(* Logix 5000 project; controller PLC_MCC1201_220AP1 vendor 1 type 14 code 164 rev 35.11; software revision 35.00; part 3 of 25 *)

   M212_M1_DR_MSF : MOTION_INSTRUCTION := (FLAGS := 570425344, DN := 1, STATUS := 2, STATE := 1); {access None}
   M212_M1_DR_MSO : MOTION_INSTRUCTION := (FLAGS := -1610612736, EN := 1, DN := 1, STATE := 1); {access None}
   M212_M1_DR_OUT_MAJ : MOTION_INSTRUCTION := (FLAGS := 570425344, DN := 1); {access None}
   M212_M1_DR_OUT_MAM : MOTION_INSTRUCTION := (FLAGS := 33554432); {access None}
   M212_M1_DR_OUT_MAR : MOTION_INSTRUCTION := (FLAGS := 33554432); {access None}
   M212_M1_DR_OUT_MAS : MOTION_INSTRUCTION := (FLAGS := -1442840576, EN := 1, DN := 1, PC := 1); {access None}
   M212_M1_DR_OUT_MCD : MOTION_INSTRUCTION := (FLAGS := 570425344, DN := 1); {access None}
   M212_M1_DR_OUT_MRP : MOTION_INSTRUCTION := (FLAGS := 33554432); {access None}
   M213_M1_DR : AXIS_CIP_DRIVE; {access Read Only}
   M213_M1_DR_IN_MAJ : MOTION_INSTRUCTION := (FLAGS := 570425344, DN := 1); {access None}
   M213_M1_DR_IN_MAM : MOTION_INSTRUCTION := (FLAGS := 33554432); {access None}
   M213_M1_DR_IN_MAR : MOTION_INSTRUCTION := (FLAGS := 33554432); {access None}
   M213_M1_DR_IN_MAS : MOTION_INSTRUCTION := (FLAGS := -1442840576, EN := 1, DN := 1, PC := 1); {access None}
   M213_M1_DR_IN_MCD : MOTION_INSTRUCTION := (FLAGS := 570425344, DN := 1); {access None}
   M213_M1_DR_IN_MRP : MOTION_INSTRUCTION := (FLAGS := 33554432); {access None}
   M213_M1_DR_MAFR : MOTION_INSTRUCTION := (FLAGS := 301989888, ER := 1, ERR := 11); {access None}
   M213_M1_DR_MDR : MOTION_INSTRUCTION := (FLAGS := -1845493760, EN := 1, ER := 1, ERR := 11); {access None}
   M213_M1_DR_MSF : MOTION_INSTRUCTION := (FLAGS := 570425344, DN := 1, STATUS := 2, STATE := 1); {access None}
   M213_M1_DR_MSO : MOTION_INSTRUCTION := (FLAGS := -1610612736, EN := 1, DN := 1, STATE := 1); {access None}
   M213_M1_DR_OUT_MAJ : MOTION_INSTRUCTION := (FLAGS := 570425344, DN := 1); {access None}
   M213_M1_DR_OUT_MAM : MOTION_INSTRUCTION := (FLAGS := 33554432); {access None}
   M213_M1_DR_OUT_MAR : MOTION_INSTRUCTION := (FLAGS := 33554432); {access None}
   M213_M1_DR_OUT_MAS : MOTION_INSTRUCTION := (FLAGS := -1442840576, EN := 1, DN := 1, PC := 1); {access None}
   M213_M1_DR_OUT_MCD : MOTION_INSTRUCTION := (FLAGS := 570425344, DN := 1); {access None}
   M213_M1_DR_OUT_MRP : MOTION_INSTRUCTION := (FLAGS := 33554432); {access None}
   M213A_M1_DR_IN_MAJ : MOTION_INSTRUCTION := (FLAGS := 570425344, DN := 1); {access None}
   M213A_M1_DR_IN_MAM : MOTION_INSTRUCTION := (FLAGS := 33554432); {access None}
   M213A_M1_DR_IN_MAR : MOTION_INSTRUCTION := (FLAGS := 33554432); {access None}
   M213A_M1_DR_IN_MAS : MOTION_INSTRUCTION := (FLAGS := -1442840576, EN := 1, DN := 1, PC := 1); {access None}
   M213A_M1_DR_IN_MCD : MOTION_INSTRUCTION := (FLAGS := 570425344, DN := 1); {access None}
   M213A_M1_DR_IN_MRP : MOTION_INSTRUCTION := (FLAGS := 33554432); {access None}
   M213A_M1_DR_MAFR : MOTION_INSTRUCTION := (FLAGS := 301989888, ER := 1, ERR := 11); {access None}
   M213A_M1_DR_MDR : MOTION_INSTRUCTION := (FLAGS := -1845493760, EN := 1, ER := 1, ERR := 11); {access None}
   M213A_M1_DR_MSF : MOTION_INSTRUCTION := (FLAGS := 570425344, DN := 1, STATUS := 2, STATE := 1); {access None}
   M213A_M1_DR_MSO : MOTION_INSTRUCTION := (FLAGS := -1610612736, EN := 1, DN := 1, STATE := 1); {access None}
   M213A_M1_DR_OUT_MAJ : MOTION_INSTRUCTION := (FLAGS := 570425344, DN := 1); {access None}
   M213A_M1_DR_OUT_MAM : MOTION_INSTRUCTION := (FLAGS := 33554432); {access None}
   M213A_M1_DR_OUT_MAR : MOTION_INSTRUCTION := (FLAGS := 33554432); {access None}
   M213A_M1_DR_OUT_MAS : MOTION_INSTRUCTION := (FLAGS := -1442840576, EN := 1, DN := 1, PC := 1); {access None}
   M213A_M1_DR_OUT_MCD : MOTION_INSTRUCTION := (FLAGS := 570425344, DN := 1); {access None}
   M213A_M1_DR_OUT_MRP : MOTION_INSTRUCTION := (FLAGS := 33554432); {access None}
   M213B_M1_DR_IN_MAJ : MOTION_INSTRUCTION := (FLAGS := 570425344, DN := 1); {access None}
   M213B_M1_DR_IN_MAM : MOTION_INSTRUCTION := (FLAGS := 33554432); {access None}
   M213B_M1_DR_IN_MAR : MOTION_INSTRUCTION := (FLAGS := 33554432); {access None}
   M213B_M1_DR_IN_MAS : MOTION_INSTRUCTION := (FLAGS := -1442840576, EN := 1, DN := 1, PC := 1); {access None}
   M213B_M1_DR_IN_MCD : MOTION_INSTRUCTION := (FLAGS := 570425344, DN := 1); {access None}
   M213B_M1_DR_IN_MRP : MOTION_INSTRUCTION := (FLAGS := 33554432); {access None}
   M213B_M1_DR_MAFR : MOTION_INSTRUCTION := (FLAGS := 301989888, ER := 1, ERR := 11); {access None}
   M213B_M1_DR_MDR : MOTION_INSTRUCTION := (FLAGS := -1845493760, EN := 1, ER := 1, ERR := 11); {access None}
   M213B_M1_DR_MSF : MOTION_INSTRUCTION := (FLAGS := 570425344, DN := 1, STATUS := 2, STATE := 1); {access None}
   M213B_M1_DR_MSO : MOTION_INSTRUCTION := (FLAGS := -1610612736, EN := 1, DN := 1, STATE := 1); {access None}
   M213B_M1_DR_OUT_MAJ : MOTION_INSTRUCTION := (FLAGS := 570425344, DN := 1); {access None}
   M213B_M1_DR_OUT_MAM : MOTION_INSTRUCTION := (FLAGS := 33554432); {access None}
   M213B_M1_DR_OUT_MAR : MOTION_INSTRUCTION := (FLAGS := 33554432); {access None}
   M213B_M1_DR_OUT_MAS : MOTION_INSTRUCTION := (FLAGS := -1442840576, EN := 1, DN := 1, PC := 1); {access None}
   M213B_M1_DR_OUT_MCD : MOTION_INSTRUCTION := (FLAGS := 570425344, DN := 1); {access None}
   M213B_M1_DR_OUT_MRP : MOTION_INSTRUCTION := (FLAGS := 33554432); {access None}
   M214_M1_DR : AXIS_CIP_DRIVE; {access Read Only}
   M214_M1_DR_IN_MAJ : MOTION_INSTRUCTION := (FLAGS := 570425344, DN := 1); {access None}
   M214_M1_DR_IN_MAM : MOTION_INSTRUCTION := (FLAGS := 33554432); {access None}
   M214_M1_DR_IN_MAR : MOTION_INSTRUCTION := (FLAGS := 33554432); {access None}
   M214_M1_DR_IN_MAS : MOTION_INSTRUCTION := (FLAGS := -1442840576, EN := 1, DN := 1, PC := 1); {access None}
   M214_M1_DR_IN_MCD : MOTION_INSTRUCTION := (FLAGS := 570425344, DN := 1); {access None}
   M214_M1_DR_IN_MRP : MOTION_INSTRUCTION := (FLAGS := 33554432); {access None}
   M214_M1_DR_MAFR : MOTION_INSTRUCTION := (FLAGS := 301989888, ER := 1, ERR := 11); {access None}
   M214_M1_DR_MDR : MOTION_INSTRUCTION := (FLAGS := -1845493760, EN := 1, ER := 1, ERR := 11); {access None}
   M214_M1_DR_MSF : MOTION_INSTRUCTION := (FLAGS := 570425344, DN := 1, STATUS := 2, STATE := 1); {access None}
   M214_M1_DR_MSO : MOTION_INSTRUCTION := (FLAGS := -1610612736, EN := 1, DN := 1, STATE := 1); {access None}
   M214_M1_DR_OUT_MAJ : MOTION_INSTRUCTION := (FLAGS := 570425344, DN := 1); {access None}
   M214_M1_DR_OUT_MAM : MOTION_INSTRUCTION := (FLAGS := 33554432); {access None}
   M214_M1_DR_OUT_MAR : MOTION_INSTRUCTION := (FLAGS := 33554432); {access None}
   M214_M1_DR_OUT_MAS : MOTION_INSTRUCTION := (FLAGS := -1442840576, EN := 1, DN := 1, PC := 1); {access None}
   M214_M1_DR_OUT_MCD : MOTION_INSTRUCTION := (FLAGS := 570425344, DN := 1); {access None}
   M214_M1_DR_OUT_MRP : MOTION_INSTRUCTION := (FLAGS := 33554432); {access None}
   M215_M1_DR : AXIS_CIP_DRIVE; {access Read Only}
   M215_M1_DR_IN_MAJ : MOTION_INSTRUCTION := (FLAGS := 570425344, DN := 1); {access None}
   M215_M1_DR_IN_MAM : MOTION_INSTRUCTION := (FLAGS := 33554432); {access None}
   M215_M1_DR_IN_MAR : MOTION_INSTRUCTION := (FLAGS := 33554432); {access None}
   M215_M1_DR_IN_MAS : MOTION_INSTRUCTION := (FLAGS := -1442840576, EN := 1, DN := 1, PC := 1); {access None}
   M215_M1_DR_IN_MCD : MOTION_INSTRUCTION := (FLAGS := 570425344, DN := 1); {access None}
   M215_M1_DR_IN_MRP : MOTION_INSTRUCTION := (FLAGS := 33554432); {access None}
   M215_M1_DR_MAFR : MOTION_INSTRUCTION := (FLAGS := 301989888, ER := 1, ERR := 11); {access None}
   M215_M1_DR_MDR : MOTION_INSTRUCTION := (FLAGS := -1845493760, EN := 1, ER := 1, ERR := 11); {access None}
   M215_M1_DR_MSF : MOTION_INSTRUCTION := (FLAGS := 570425344, DN := 1, STATUS := 2, STATE := 1); {access None}
   M215_M1_DR_MSO : MOTION_INSTRUCTION := (FLAGS := -1610612736, EN := 1, DN := 1, STATE := 1); {access None}
   M215_M1_DR_OUT_MAJ : MOTION_INSTRUCTION := (FLAGS := 570425344, DN := 1); {access None}
   M215_M1_DR_OUT_MAM : MOTION_INSTRUCTION := (FLAGS := 33554432); {access None}
   M215_M1_DR_OUT_MAR : MOTION_INSTRUCTION := (FLAGS := 33554432); {access None}
   M215_M1_DR_OUT_MAS : MOTION_INSTRUCTION := (FLAGS := -1442840576, EN := 1, DN := 1, PC := 1); {access None}
   M215_M1_DR_OUT_MCD : MOTION_INSTRUCTION := (FLAGS := 570425344, DN := 1); {access None}
   M215_M1_DR_OUT_MRP : MOTION_INSTRUCTION := (FLAGS := 33554432); {access None}
   M216_M1_DR : AXIS_CIP_DRIVE; {access Read Only}
   M216_M1_DR_IN_MAJ : MOTION_INSTRUCTION := (FLAGS := 570425344, DN := 1); {access None}
   M216_M1_DR_IN_MAM : MOTION_INSTRUCTION := (FLAGS := 33554432); {access None}
   M216_M1_DR_IN_MAR : MOTION_INSTRUCTION := (FLAGS := 33554432); {access None}
   M216_M1_DR_IN_MAS : MOTION_INSTRUCTION := (FLAGS := -1442840576, EN := 1, DN := 1, PC := 1); {access None}
   M216_M1_DR_IN_MCD : MOTION_INSTRUCTION := (FLAGS := 570425344, DN := 1); {access None}
   M216_M1_DR_IN_MRP : MOTION_INSTRUCTION := (FLAGS := 33554432); {access None}
   M216_M1_DR_MAFR : MOTION_INSTRUCTION := (FLAGS := 301989888, ER := 1, ERR := 11); {access None}
   M216_M1_DR_MDR : MOTION_INSTRUCTION := (FLAGS := -1845493760, EN := 1, ER := 1, ERR := 11); {access None}
   M216_M1_DR_MSF : MOTION_INSTRUCTION := (FLAGS := 570425344, DN := 1, STATUS := 2, STATE := 1); {access None}
   M216_M1_DR_MSO : MOTION_INSTRUCTION := (FLAGS := -1610612736, EN := 1, DN := 1, STATE := 1); {access None}
   M216_M1_DR_OUT_MAJ : MOTION_INSTRUCTION := (FLAGS := 570425344, DN := 1); {access None}
   M216_M1_DR_OUT_MAM : MOTION_INSTRUCTION := (FLAGS := 33554432); {access None}
   M216_M1_DR_OUT_MAR : MOTION_INSTRUCTION := (FLAGS := 33554432); {access None}
   M216_M1_DR_OUT_MAS : MOTION_INSTRUCTION := (FLAGS := -1442840576, EN := 1, DN := 1, PC := 1); {access None}
   M216_M1_DR_OUT_MCD : MOTION_INSTRUCTION := (FLAGS := 570425344, DN := 1); {access None}
   M216_M1_DR_OUT_MRP : MOTION_INSTRUCTION := (FLAGS := 33554432); {access None}
   M217_M1_DR : AXIS_CIP_DRIVE; {access Read Only}
   M217_M1_DR_IN_MAJ : MOTION_INSTRUCTION := (FLAGS := 570425344, DN := 1); {access None}
   M217_M1_DR_IN_MAM : MOTION_INSTRUCTION := (FLAGS := 33554432); {access None}
   M217_M1_DR_IN_MAR : MOTION_INSTRUCTION := (FLAGS := 33554432); {access None}
   M217_M1_DR_IN_MAS : MOTION_INSTRUCTION := (FLAGS := -1442840576, EN := 1, DN := 1, PC := 1); {access None}
   M217_M1_DR_IN_MCD : MOTION_INSTRUCTION := (FLAGS := 570425344, DN := 1); {access None}
   M217_M1_DR_IN_MRP : MOTION_INSTRUCTION := (FLAGS := 33554432); {access None}
   M217_M1_DR_MAFR : MOTION_INSTRUCTION := (FLAGS := 301989888, ER := 1, ERR := 11); {access None}
   M217_M1_DR_MDR : MOTION_INSTRUCTION := (FLAGS := -1845493760, EN := 1, ER := 1, ERR := 11); {access None}
   M217_M1_DR_MSF : MOTION_INSTRUCTION := (FLAGS := 570425344, DN := 1, STATUS := 2, STATE := 1); {access None}
   M217_M1_DR_MSO : MOTION_INSTRUCTION := (FLAGS := -1610612736, EN := 1, DN := 1, STATE := 1); {access None}
   M217_M1_DR_OUT_MAJ : MOTION_INSTRUCTION := (FLAGS := 570425344, DN := 1); {access None}
   M217_M1_DR_OUT_MAM : MOTION_INSTRUCTION := (FLAGS := 33554432); {access None}
   M217_M1_DR_OUT_MAR : MOTION_INSTRUCTION := (FLAGS := 33554432); {access None}
   M217_M1_DR_OUT_MAS : MOTION_INSTRUCTION := (FLAGS := -1442840576, EN := 1, DN := 1, PC := 1); {access None}
   M217_M1_DR_OUT_MCD : MOTION_INSTRUCTION := (FLAGS := 570425344, DN := 1); {access None}
   M217_M1_DR_OUT_MRP : MOTION_INSTRUCTION := (FLAGS := 33554432); {access None}
   M218_M1_DR : AXIS_CIP_DRIVE; {access Read Only}
   M218_M1_DR_IN_MAJ : MOTION_INSTRUCTION := (FLAGS := 570425344, DN := 1); {access None}
   M218_M1_DR_IN_MAM : MOTION_INSTRUCTION := (FLAGS := 33554432); {access None}
   M218_M1_DR_IN_MAR : MOTION_INSTRUCTION := (FLAGS := 33554432); {access None}
   M218_M1_DR_IN_MAS : MOTION_INSTRUCTION := (FLAGS := -1442840576, EN := 1, DN := 1, PC := 1); {access None}
   M218_M1_DR_IN_MCD : MOTION_INSTRUCTION := (FLAGS := 570425344, DN := 1); {access None}
   M218_M1_DR_IN_MRP : MOTION_INSTRUCTION := (FLAGS := 33554432); {access None}
   M218_M1_DR_MAFR : MOTION_INSTRUCTION := (FLAGS := 301989888, ER := 1, ERR := 11); {access None}
   M218_M1_DR_MDR : MOTION_INSTRUCTION := (FLAGS := -1845493760, EN := 1, ER := 1, ERR := 11); {access None}
   M218_M1_DR_MSF : MOTION_INSTRUCTION := (FLAGS := 570425344, DN := 1, STATUS := 2, STATE := 1); {access None}
   M218_M1_DR_MSO : MOTION_INSTRUCTION := (FLAGS := -1610612736, EN := 1, DN := 1, STATE := 1); {access None}
   M218_M1_DR_OUT_MAJ : MOTION_INSTRUCTION := (FLAGS := 570425344, DN := 1); {access None}
   M218_M1_DR_OUT_MAM : MOTION_INSTRUCTION := (FLAGS := 33554432); {access None}
   M218_M1_DR_OUT_MAR : MOTION_INSTRUCTION := (FLAGS := 33554432); {access None}
   M218_M1_DR_OUT_MAS : MOTION_INSTRUCTION := (FLAGS := -1442840576, EN := 1, DN := 1, PC := 1); {access None}
   M218_M1_DR_OUT_MCD : MOTION_INSTRUCTION := (FLAGS := 570425344, DN := 1); {access None}
   M218_M1_DR_OUT_MRP : MOTION_INSTRUCTION := (FLAGS := 33554432); {access None}
   M219_M1_DR : AXIS_CIP_DRIVE; {access Read Only}
   M219_M1_DR_IN_MAJ : MOTION_INSTRUCTION := (FLAGS := 570425344, DN := 1); {access None}
   M219_M1_DR_IN_MAM : MOTION_INSTRUCTION := (FLAGS := 33554432); {access None}
   M219_M1_DR_IN_MAR : MOTION_INSTRUCTION := (FLAGS := 33554432); {access None}
   M219_M1_DR_IN_MAS : MOTION_INSTRUCTION := (FLAGS := -1442840576, EN := 1, DN := 1, PC := 1); {access None}
   M219_M1_DR_IN_MCD : MOTION_INSTRUCTION := (FLAGS := 570425344, DN := 1); {access None}
   M219_M1_DR_IN_MRP : MOTION_INSTRUCTION := (FLAGS := 33554432); {access None}
   M219_M1_DR_MAFR : MOTION_INSTRUCTION := (FLAGS := 301989888, ER := 1, ERR := 11); {access None}
   M219_M1_DR_MDR : MOTION_INSTRUCTION := (FLAGS := -1845493760, EN := 1, ER := 1, ERR := 11); {access None}
   M219_M1_DR_MSF : MOTION_INSTRUCTION := (FLAGS := 570425344, DN := 1, STATUS := 2, STATE := 1); {access None}
   M219_M1_DR_MSO : MOTION_INSTRUCTION := (FLAGS := -1610612736, EN := 1, DN := 1, STATE := 1); {access None}
   M219_M1_DR_OUT_MAJ : MOTION_INSTRUCTION := (FLAGS := 570425344, DN := 1); {access None}
   M219_M1_DR_OUT_MAM : MOTION_INSTRUCTION := (FLAGS := 33554432); {access None}
   M219_M1_DR_OUT_MAR : MOTION_INSTRUCTION := (FLAGS := 33554432); {access None}
   M219_M1_DR_OUT_MAS : MOTION_INSTRUCTION := (FLAGS := -1442840576, EN := 1, DN := 1, PC := 1); {access None}
   M219_M1_DR_OUT_MCD : MOTION_INSTRUCTION := (FLAGS := 570425344, DN := 1); {access None}
   M219_M1_DR_OUT_MRP : MOTION_INSTRUCTION := (FLAGS := 33554432); {access None}
   M220_M1_DR : AXIS_CIP_DRIVE; {access Read Only}
   M220_M1_DR_IN_MAJ : MOTION_INSTRUCTION := (FLAGS := 570425344, DN := 1); {access None}
   M220_M1_DR_IN_MAM : MOTION_INSTRUCTION := (FLAGS := 33554432); {access None}
   M220_M1_DR_IN_MAR : MOTION_INSTRUCTION := (FLAGS := 33554432); {access None}
   M220_M1_DR_IN_MAS : MOTION_INSTRUCTION := (FLAGS := -1442840576, EN := 1, DN := 1, PC := 1); {access None}
   M220_M1_DR_IN_MCD : MOTION_INSTRUCTION := (FLAGS := 570425344, DN := 1); {access None}
   M220_M1_DR_IN_MRP : MOTION_INSTRUCTION := (FLAGS := 33554432); {access None}
   M220_M1_DR_MAFR : MOTION_INSTRUCTION := (FLAGS := 301989888, ER := 1, ERR := 11); {access None}
   M220_M1_DR_MDR : MOTION_INSTRUCTION := (FLAGS := -1845493760, EN := 1, ER := 1, ERR := 11); {access None}
   M220_M1_DR_MSF : MOTION_INSTRUCTION := (FLAGS := 570425344, DN := 1, STATUS := 2, STATE := 1); {access None}
   M220_M1_DR_MSO : MOTION_INSTRUCTION := (FLAGS := -1610612736, EN := 1, DN := 1, STATE := 1); {access None}
   M220_M1_DR_OUT_MAJ : MOTION_INSTRUCTION := (FLAGS := 570425344, DN := 1); {access None}
   M220_M1_DR_OUT_MAM : MOTION_INSTRUCTION := (FLAGS := 33554432); {access None}
   M220_M1_DR_OUT_MAR : MOTION_INSTRUCTION := (FLAGS := 33554432); {access None}
   M220_M1_DR_OUT_MAS : MOTION_INSTRUCTION := (FLAGS := -1442840576, EN := 1, DN := 1, PC := 1); {access None}
   M220_M1_DR_OUT_MCD : MOTION_INSTRUCTION := (FLAGS := 570425344, DN := 1); {access None}
   M220_M1_DR_OUT_MRP : MOTION_INSTRUCTION := (FLAGS := 33554432); {access None}
   M225 : MAC_EMERGENCYXCUT := (ST_xConditionOKAccessArea := 1, ST_xSelectorManualMode := 1, ST_xManualModeSelection := 1, ST_xManualModeAccepted := 1, ST_xDistanceBetweenCutOK := 1, ST_xConditionOKStopCycle := 1, ST_xConditionOKSemiautoMode := 1, ST_xConditionOKManualMode := 1, ST_xBreakerCutRequest := 1, OUTPUT_xMachineOutOfOrder := 1, OUTPUT_xAreaSafetyOn := 1, OUTPUT_xStopCut := 1, AUX_dDistanceFTCHead := 6050, AUX_dBridgeAngle := 80000, AUX_dManualSpeed_mm_min := 10000, AUX_dRiseReactionTime_ms := 50, AUX_dDescentReactionTime_ms := 1000, AUX_dBackwardFastSpeed_mm_min := 120000, AUX_dBackwardSlowSpeed_mm_min := 90000, AUX_dCarriageFinalPosition_cmm := 400000, AUX_dMinimumStripeLength := 100000, AUX_dMaximumStripeLength := 300000, AUX_dLastCutValue := -268936272, AUX_dLastCutValueStored := -268936272, AUX_dForwardTimeoutTime_ms := 2147483647, AUX_dReturnSpeed_mm_min := 90000, AUX_dReqSpeed_mm_min := 10000, AUX_dStartControlPhotocellPos_dmm := -36050, AUX_dTimeFTCToHead_ms := 36300000, AUX_dTimeDelayToDescent_ms := 36299800, AUX_dTimeAdvanceToRise_ms := 36293450, AUX_dTimeDelayToLubrication_ms := 36300000, OSR_xConditionNotOKToCut := 1, AUX_tmOFF_DriveEnable.PRE := 100, AUX_tmOFF_DriveEnable.ACC := 100, AUX_tmOFF_AreaSafetyOK.PRE := 2000, AUX_tmOFF_AreaSafetyOK.ACC := 2000, AUX_tmON_FdbkError.PRE := 2000, AUX_tmON_TimeoutHome.PRE := 90000, AUX_tmON_TimeoutFW.PRE := 120000, AUX_tmON_TimeoutBW.PRE := 90000, AUX_tmOFF_LowerHeadNotAllowed.PRE := 200, AUX_tmOFF_LowerHeadNotAllowed.ACC := 200, AUX_tmOFF_AdvanceTimeToRise.PRE := 171, AUX_tmOFF_AdvanceTimeToRise.ACC := 171, AUX_tmON_DelayTimeLubrication.PRE := 221, AUX_tmON_DelayTimeLubrication.ACC := 221, AUX_tmON_TimeoutHeadPosition.PRE := 90000, CONST_dAcceleration_m_s2 := 3, CONST_dDeceleration_m_s2 := 3); {access None}
   M225_ALM : MAC_EMERGENCYXCUT_ALM; {access Read Only}
        .rgxStoppingFaults[0].4   // A120KE1.Area safety
        .rgxStoppingFaults[0].8   // A57AZ1.Timeout move backward
        .rgxStoppingFaults[0].2   // A57AZ1.Drive error
        .rgxStoppingFaults[0].9   // A57AZ1.Timeout home position (A121SQ1)
        .rgxStoppingFaults[0].1   // A207BT2.Motor thermal probe
        .rgxFaults[0].0   // A57QM1.Protection traslation
        .rgxFaults[0].1   // A57QM2.Protection fan rotation
        .rgdCodeAlarm[0].0   // A63AZ1.Code alarm
        .rgxStoppingFaults[0].7   // A57AZ1.Timeout move forward
        .rgxStoppingFaults[0].11   // A207SP1.Compressed air failure
        .rgxStoppingFaults[0].10   // A208SQ1.Error position cutting head
        .rgxStoppingFaults[0].5   // A121SQ1.Forward Overstroke
        .rgxStoppingFaults[0].6   // A121SQ2.Backward Overstroke
        .rgxStoppingFaults[0].3   // A57AZ1.Traslation feedback
        .rgxStoppingFaults[0].0   // A57QS1.Safety motor sectioning
   M225_HMR : MAC_EMERGENCYXCUT_HMR := (dMode := 1, dStatus := 1, dZoneStatus := 2, dDistanceFromSnaproll_cmm := 5050000, rHeadUsage_km := 0.0004); {access Read Only}
   M225_HMW : MAC_EMERGENCYXCUT_HMW := (dLowerHeadDelayTime_ms := 800, dRiseHeadAdvanceTime_ms := 6500, dCulletStripeLength_cmm := 220000, dDistanceFromSnaproll_cmm := 5030000);
   M225_IN_MOTION : MAC_EMERGENCYXCUT_IN_MOTION; {access None}
   M225_M1_DR : AXIS_CIP_DRIVE; {access Read Only}
   M225_M1_DR_IN_MAJ : MOTION_INSTRUCTION := (FLAGS := 570425344, DN := 1); {access None}
   M225_M1_DR_IN_MAM : MOTION_INSTRUCTION := (FLAGS := 33554432); {access None}
   M225_M1_DR_IN_MAR : MOTION_INSTRUCTION := (FLAGS := 33554432); {access None}
   M225_M1_DR_IN_MAS : MOTION_INSTRUCTION := (FLAGS := -1442840576, EN := 1, DN := 1, PC := 1); {access None}
   M225_M1_DR_IN_MCD : MOTION_INSTRUCTION := (FLAGS := 570425344, DN := 1); {access None}
   M225_M1_DR_IN_MRP : MOTION_INSTRUCTION := (FLAGS := 33554432); {access None}
   M225_M1_DR_MAFR : MOTION_INSTRUCTION := (FLAGS := 301989888, ER := 1, ERR := 11); {access None}
   M225_M1_DR_MDR : MOTION_INSTRUCTION := (FLAGS := -1845493760, EN := 1, ER := 1, ERR := 11); {access None}
   M225_M1_DR_MSF : MOTION_INSTRUCTION := (FLAGS := 570425344, DN := 1, STATUS := 2, STATE := 1); {access None}
   M225_M1_DR_MSO : MOTION_INSTRUCTION := (FLAGS := -1610612736, EN := 1, DN := 1, STATE := 1); {access None}
   M225_M1_DR_OUT_MAJ : MOTION_INSTRUCTION := (FLAGS := 570425344, DN := 1); {access None}
   M225_M1_DR_OUT_MAM : MOTION_INSTRUCTION := (FLAGS := 33554432); {access None}
   M225_M1_DR_OUT_MAR : MOTION_INSTRUCTION := (FLAGS := 33554432); {access None}
   M225_M1_DR_OUT_MAS : MOTION_INSTRUCTION := (FLAGS := -1442840576, EN := 1, DN := 1, PC := 1); {access None}
   M225_M1_DR_OUT_MCD : MOTION_INSTRUCTION := (FLAGS := 570425344, DN := 1); {access None}
   M225_M1_DR_OUT_MRP : MOTION_INSTRUCTION := (FLAGS := 33554432); {access None}
   M225_OUT_MOTION : MAC_EMERGENCYXCUT_OUT_MOTION := (DR_MSO.FLAGS := 33554432, DR_MSF.FLAGS := -1577058304, DR_MSF.EN := 1, DR_MSF.DN := 1, DR_MSF.STATUS := 2, DR_MSF.STATE := 1, DR_MASR.FLAGS := 33554432, DR_MAJ.FLAGS := 33554432, DR_MAM.FLAGS := 33554432, DR_MAS.FLAGS := -1442840576, DR_MAS.EN := 1, DR_MAS.DN := 1, DR_MAS.PC := 1, DR_MAH.FLAGS := 33554432); {access None}
   M225S_AOI_AccessArea : STRUCT_AccessArea := (tAccess[0].tHMR.dStatusAccessArea := 4, tAccess[0].tSTC.IN_xConditionOkAccessArea := 1, tAccess[0].tSTC.OUT_xSafetyAreaIntervened := 1, tAccess[1].tHMR.dStatusAccessArea := 4, tAccess[1].tSTC.OUT_xSafetyAreaIntervened := 1);
   M2xx_CONVEYOR : MAC_CONVEYOR[20] := ([0].AUX_tmOFFRetainDriveEnable.PRE := 1000, [0].AUX_tmOFFRetainDriveEnable.ACC := 1000, [0].AUX_tmONRotfeedBackAlarm.PRE := 2000, [0].AUX_tmONDriveReadyAlarm.PRE := 1000, [0].AUX_rAcceleration_m_s2 := 0.25, [0].AUX_rDeceleration_m_s2 := 0.25, [0].AUX_dReqSpeed_mm_min := 6807, [0].AUX_dRealSpeed_mm_min := 6807, [1].AUX_tmOFFRetainDriveEnable.PRE := 1000, [1].AUX_tmOFFRetainDriveEnable.ACC := 1000, [1].AUX_tmONDriveReadyAlarm.PRE := 1000, [1].AUX_rAcceleration_m_s2 := 0.25, [1].AUX_rDeceleration_m_s2 := 0.25, [1].AUX_dReqSpeed_mm_min := 6807, [1].AUX_dRealSpeed_mm_min := 6807, [2].INPUT_xProtectionFan := 1, [2].AUX_tmOFFRetainDriveEnable.PRE := 1000, [2].AUX_tmOFFRetainDriveEnable.ACC := 1000, [2].AUX_tmONDriveReadyAlarm.PRE := 1000, [2].AUX_rAcceleration_m_s2 := 0.25, [2].AUX_rDeceleration_m_s2 := 0.25, [2].AUX_dReqSpeed_mm_min := 6807, [2].AUX_dRealSpeed_mm_min := 6807, [3].INPUT_xProtectionFan := 1, [3].AUX_tmOFFRetainDriveEnable.PRE := 1000, [3].AUX_tmOFFRetainDriveEnable.ACC := 1000, [3].AUX_tmONDriveReadyAlarm.PRE := 1000, [3].AUX_rAcceleration_m_s2 := 0.25, [3].AUX_rDeceleration_m_s2 := 0.25, [3].AUX_dReqSpeed_mm_min := 6807, [3].AUX_dRealSpeed_mm_min := 6807, [4].INPUT_xProtectionFan := 1, [4].AUX_tmOFFRetainDriveEnable.PRE := 1000, [4].AUX_tmOFFRetainDriveEnable.ACC := 1000, [4].AUX_tmONDriveReadyAlarm.PRE := 1000, [4].AUX_rAcceleration_m_s2 := 0.25, [4].AUX_rDeceleration_m_s2 := 0.25, [4].AUX_dReqSpeed_mm_min := 6807, [4].AUX_dRealSpeed_mm_min := 6807, [5].ST_xStoppingFaults := 1, [5].INPUT_xProtectionFan := 1, [5].AUX_tmOFFRetainDriveEnable.PRE := 1000, [5].AUX_tmOFFRetainDriveEnable.ACC := 1000, [5].AUX_tmONDriveReadyAlarm.PRE := 1000, [5].AUX_rAcceleration_m_s2 := 0.25, [5].AUX_rDeceleration_m_s2 := 0.25, [5].AUX_dReqSpeed_mm_min := 6807, [5].AUX_dRealSpeed_mm_min := 6807, [6].ST_xStoppingFaults := 1, [6].INPUT_xProtectionFan := 1, [6].AUX_tmOFFRetainDriveEnable.PRE := 1000, [6].AUX_tmOFFRetainDriveEnable.ACC := 1000, [6].AUX_tmONDriveReadyAlarm.PRE := 1000, [6].AUX_rAcceleration_m_s2 := 0.25, [6].AUX_rDeceleration_m_s2 := 0.25, [6].AUX_dReqSpeed_mm_min := 6807, [6].AUX_dRealSpeed_mm_min := 6807, [7].ST_xStoppingFaults := 1, [7].INPUT_xProtectionFan := 1, [7].AUX_tmOFFRetainDriveEnable.PRE := 1000,
        [7].AUX_tmOFFRetainDriveEnable.ACC := 1000, [7].AUX_tmONDriveReadyAlarm.PRE := 1000, [7].AUX_rAcceleration_m_s2 := 0.25, [7].AUX_rDeceleration_m_s2 := 0.25, [7].AUX_dReqSpeed_mm_min := 6807, [7].AUX_dRealSpeed_mm_min := 6807, [8].ST_xStoppingFaults := 1, [8].INPUT_xProtectionFan := 1, [8].AUX_tmOFFRetainDriveEnable.PRE := 1000, [8].AUX_tmOFFRetainDriveEnable.ACC := 1000, [8].AUX_tmONDriveReadyAlarm.PRE := 1000, [8].AUX_rAcceleration_m_s2 := 0.25, [8].AUX_rDeceleration_m_s2 := 0.25, [8].AUX_dReqSpeed_mm_min := 6807, [8].AUX_dRealSpeed_mm_min := 6807, [9].ST_xStoppingFaults := 1, [9].INPUT_xProtectionFan := 1, [9].AUX_tmOFFRetainDriveEnable.PRE := 1000, [9].AUX_tmOFFRetainDriveEnable.ACC := 1000, [9].AUX_tmONDriveReadyAlarm.PRE := 1000, [9].AUX_rAcceleration_m_s2 := 0.25, [9].AUX_rDeceleration_m_s2 := 0.25, [9].AUX_dReqSpeed_mm_min := 6807, [9].AUX_dRealSpeed_mm_min := 6807, [10].ST_xStoppingFaults := 1, [10].INPUT_xProtectionFan := 1, [10].AUX_tmOFFRetainDriveEnable.PRE := 1000, [10].AUX_tmOFFRetainDriveEnable.ACC := 1000, [10].AUX_tmONDriveReadyAlarm.PRE := 1000, [10].AUX_rAcceleration_m_s2 := 0.25, [10].AUX_rDeceleration_m_s2 := 0.25, [10].AUX_dReqSpeed_mm_min := 6807, [10].AUX_dRealSpeed_mm_min := 6807, [11].INPUT_xProtectionFan := 1, [11].AUX_tmOFFRetainDriveEnable.PRE := 1000, [11].AUX_tmOFFRetainDriveEnable.ACC := 1000, [11].AUX_tmONDriveReadyAlarm.PRE := 1000, [11].AUX_rAcceleration_m_s2 := 0.25, [11].AUX_rDeceleration_m_s2 := 0.25, [11].AUX_dReqSpeed_mm_min := 6807, [11].AUX_dRealSpeed_mm_min := 6807, [12].INPUT_xProtectionFan := 1, [12].AUX_tmOFFRetainDriveEnable.PRE := 1000, [12].AUX_tmOFFRetainDriveEnable.ACC := 1000, [12].AUX_dReqSpeed_mm_min := 6807, [12].AUX_dRealSpeed_mm_min := 6807, [13].INPUT_xProtectionFan := 1, [13].AUX_tmOFFRetainDriveEnable.PRE := 1000, [13].AUX_tmOFFRetainDriveEnable.ACC := 1000, [13].AUX_dReqSpeed_mm_min := 6807, [13].AUX_dRealSpeed_mm_min := 6807, [14].INPUT_xProtectionFan := 1, [14].AUX_tmOFFRetainDriveEnable.PRE := 1000, [14].AUX_tmOFFRetainDriveEnable.ACC := 1000, [14].AUX_dReqSpeed_mm_min := 6807, [14].AUX_dRealSpeed_mm_min := 6807, [15].INPUT_xProtectionFan := 1, [15].AUX_tmOFFRetainDriveEnable.PRE := 1000, [15].AUX_tmOFFRetainDriveEnable.ACC := 1000, [15].AUX_dReqSpeed_mm_min := 6807,
        [15].AUX_dRealSpeed_mm_min := 6807, [16].INPUT_xProtectionFan := 1, [16].AUX_tmOFFRetainDriveEnable.PRE := 1000, [16].AUX_tmOFFRetainDriveEnable.ACC := 1000, [16].AUX_dReqSpeed_mm_min := 6807, [16].AUX_dRealSpeed_mm_min := 6807, [17].INPUT_xProtectionFan := 1, [17].AUX_tmOFFRetainDriveEnable.PRE := 1000, [17].AUX_tmOFFRetainDriveEnable.ACC := 1000, [17].AUX_dReqSpeed_mm_min := 6807, [17].AUX_dRealSpeed_mm_min := 6807, [18].INPUT_xProtectionFan := 1, [18].AUX_tmOFFRetainDriveEnable.PRE := 1000, [18].AUX_tmOFFRetainDriveEnable.ACC := 1000, [18].AUX_dReqSpeed_mm_min := 6807, [18].AUX_dRealSpeed_mm_min := 6807, [19].INPUT_xProtectionFan := 1, [19].AUX_tmOFFRetainDriveEnable.PRE := 1000, [19].AUX_tmOFFRetainDriveEnable.ACC := 1000, [19].AUX_dReqSpeed_mm_min := 6807, [19].AUX_dRealSpeed_mm_min := 6807); {access None}
        [0]   // M202
        [10]   // M213
        [1]   // M203
        [2]   // M204
        [3]   // M206
        [4]   // M207
        [5]   // M208
        [6]   // M209
        [7]   // M210
        [8]   // M211
        [9]   // M212
        [11]   // M214
        [12]   // M215
        [13]   // M216
        [14]   // M217
        [15]   // M218
        [19]   // M301M2
        [18]   // M301M1
        [16]   // M219
        [17]   // M220
   M2xx_CONVEYOR_ALM : MAC_CONVEYOR_ALM[20] := ([5].rgxStoppingFaults[0] := 16, [6].rgxStoppingFaults[0] := 16, [7].rgxStoppingFaults[0] := 16, [8].rgxStoppingFaults[0] := 16, [9].rgxStoppingFaults[0] := 16, [10].rgxStoppingFaults[0] := 16); {access Read Only}
        [0]   // M202
        [0].rgxStoppingFaults[0].2   // A53AZ1.Drive error
        [2].rgxStoppingFaults[0].2   // A55AZ1.Drive error
        [1].rgxStoppingFaults[0].2   // A54AZ1.Drive error
        [0].rgdCodeAlarm[0].0   // AZ.Drive error code
        [0].rgxFaults[0].0   // QM.Protection fan rotation
        [10]   // M213
        [11]   // M214
        [1]   // M203
        [2]   // M204
        [3]   // M206
        [4]   // M207
        [5]   // M208
        [6]   // M209
        [7]   // M210
        [8]   // M211
        [9]   // M212
        [17]   // M220
        [18]   // M301M1
        [16]   // M219
        [15]   // M218
        [14]   // M217
        [13]   // M216
        [12]   // M215
        [19]   // M301M2
        [0].rgxStoppingFaults[0].1   // A206BT1.Motor thermal probe
        [1].rgxStoppingFaults[0].1   // A206BT2.Motor thermal probe
        [1].rgxStoppingFaults[0].3   // A54AZ1.Rotation feedback
        [0].rgxStoppingFaults[0].0   // A53QS1.Local safety switch
        [0].rgxStoppingFaults[0].4   // A53AZ1.Drive not ready
        [1].rgxStoppingFaults[0].0   // A54QS1.Local safety switch
        [0].rgxStoppingFaults[0].3   // A53AZ1.Rotation feedback
        [1].rgxStoppingFaults[0].4   // A54AZ1.Drive not ready
        [2].rgxStoppingFaults[0].0   // A55QS1.Local safety switch
        [2].rgxStoppingFaults[0].1   // A207BT1.Motor thermal probe
        [2].rgxStoppingFaults[0].3   // A55AZ1.Rotation feedback
        [2].rgxStoppingFaults[0].4   // A55AZ1.Drive not ready
        [3].rgxStoppingFaults[0].0   // A61QS1.Local safety switch
        [3].rgxStoppingFaults[0].1   // A209BT1.Motor thermal probe
        [3].rgxStoppingFaults[0].2   // A61AZ1.Drive error
        [3].rgxStoppingFaults[0].3   // A61AZ1.Rotation feedback
        [3].rgxStoppingFaults[0].4   // A61AZ1.Drive not ready
        [4].rgxStoppingFaults[0].0   // A62QS1.Local safety switch
        [5].rgxStoppingFaults[0].0   // A63QS1.Local safety switch
        [6].rgxStoppingFaults[0].0   // A64QS1.Local safety switch
        [7].rgxStoppingFaults[0].0   // A65QS1.Local safety switch
        [8].rgxStoppingFaults[0].0   // A66QS1.Local safety switch
        [9].rgxStoppingFaults[0].0   // A67QS1.Local safety switch
        [10].rgxStoppingFaults[0].0   // A68QS1.Local safety switch
        [11].rgxStoppingFaults[0].0   // A69QS1.Local safety switch
        [12].rgxStoppingFaults[0].0   // A70QS1.Local safety switch
        [13].rgxStoppingFaults[0].0   // A71QS1.Local safety switch
        [14].rgxStoppingFaults[0].0   // A72QS1.Local safety switch
        [15].rgxStoppingFaults[0].0   // A73QS1.Local safety switch
        [16].rgxStoppingFaults[0].0   // A74QS1.Local safety switch
        [17].rgxStoppingFaults[0].0   // A77QS1.Local safety switch
        [4].rgxStoppingFaults[0].1   // A209BT2.Motor thermal probe
        [5].rgxStoppingFaults[0].1   // A209BT3.Motor thermal probe
        [6].rgxStoppingFaults[0].1   // A209BT4.Motor thermal probe
        [7].rgxStoppingFaults[0].1   // A209BT5.Motor thermal probe
        [8].rgxStoppingFaults[0].1   // A209BT6.Motor thermal probe
        [9].rgxStoppingFaults[0].1   // A209BT7.Motor thermal probe
        [10].rgxStoppingFaults[0].1   // A209BT8.Motor thermal probe
        [11].rgxStoppingFaults[0].1   // A210BT1.Motor thermal probe
        [12].rgxStoppingFaults[0].1   // A210BT2.Motor thermal probe
        [13].rgxStoppingFaults[0].1   // A210BT3.Motor thermal probe
        [14].rgxStoppingFaults[0].1   // A210BT4.Motor thermal probe
        [15].rgxStoppingFaults[0].1   // A210BT5.Motor thermal probe
        [16].rgxStoppingFaults[0].1   // A210BT6.Motor thermal probe
        [18].rgxStoppingFaults[0].1   // A210BT7.Motor thermal probe
        [19].rgxStoppingFaults[0].1   // A210BT8.Motor thermal probe
        [17].rgxStoppingFaults[0].1   // A211BT1.Motor thermal probe
        [18].rgxStoppingFaults[0].0   // A75QS1.Local safety switch
        [19].rgxStoppingFaults[0].0   // A76QS1.Local safety switch
        [4].rgxStoppingFaults[0].2   // A62AZ1.Drive error
        [4].rgxStoppingFaults[0].3   // A62AZ1.Rotation feedback
        [4].rgxStoppingFaults[0].4   // A62AZ1.Drive not ready
        [5].rgxStoppingFaults[0].2   // A63AZ1.Drive error
        [6].rgxStoppingFaults[0].2   // A64AZ1.Drive error
        [7].rgxStoppingFaults[0].2   // A65AZ1.Drive error
        [8].rgxStoppingFaults[0].2   // A66AZ1.Drive error
        [9].rgxStoppingFaults[0].2   // A67AZ1.Drive error
        [10].rgxStoppingFaults[0].2   // A68AZ1.Drive error
        [11].rgxStoppingFaults[0].2   // A69AZ1.Drive error
        [12].rgxStoppingFaults[0].2   // A70AZ1.Drive error
        [13].rgxStoppingFaults[0].2   // A71AZ1.Drive error
        [14].rgxStoppingFaults[0].2   // A72AZ1.Drive error
        [15].rgxStoppingFaults[0].2   // A73AZ1.Drive error
        [16].rgxStoppingFaults[0].2   // A74AZ1.Drive error
        [17].rgxStoppingFaults[0].2   // A77AZ1.Drive error
        [18].rgxStoppingFaults[0].2   // A75AZ1.Drive error
        [19].rgxStoppingFaults[0].2   // A76AZ1.Drive error
        [19].rgxStoppingFaults[0].3   // A76AZ1.Rotation feedback
        [18].rgxStoppingFaults[0].3   // A75AZ1.Rotation feedback
        [17].rgxStoppingFaults[0].3   // A77AZ1.Rotation feedback
        [16].rgxStoppingFaults[0].3   // A74AZ1.Rotation feedback
        [15].rgxStoppingFaults[0].3   // A73AZ1.Rotation feedback
        [14].rgxStoppingFaults[0].3   // A72AZ1.Rotation feedback
        [13].rgxStoppingFaults[0].3   // A71AZ1.Rotation feedback
        [12].rgxStoppingFaults[0].3   // A70AZ1.Rotation feedback
        [11].rgxStoppingFaults[0].3   // A69AZ1.Rotation feedback
        [10].rgxStoppingFaults[0].3   // A68AZ1.Rotation feedback
        [9].rgxStoppingFaults[0].3   // A67AZ1.Rotation feedback
        [8].rgxStoppingFaults[0].3   // A66AZ1.Rotation feedback
        [7].rgxStoppingFaults[0].3   // A65AZ1.Rotation feedback
        [6].rgxStoppingFaults[0].3   // A64AZ1.Rotation feedback
        [5].rgxStoppingFaults[0].3   // A63AZ1.Rotation feedback
        [4].rgxStoppingFaults[0].5   // A62AZ1.Rotation feedback
        [3].rgxStoppingFaults[0].5   // A61AZ1.Rotation feedback
        [3].rgxStoppingFaults[0].6   // A61AZ1.Drive not ready
        [4].rgxStoppingFaults[0].6   // A62AZ1.Drive not ready
        [5].rgxStoppingFaults[0].4   // A63AZ1.Drive not ready
        [6].rgxStoppingFaults[0].4   // A64AZ1.Drive not ready
        [7].rgxStoppingFaults[0].4   // A65AZ1.Drive not ready
        [8].rgxStoppingFaults[0].4   // A66AZ1.Drive not ready
        [9].rgxStoppingFaults[0].4   // A67AZ1.Drive not ready
        [10].rgxStoppingFaults[0].4   // A68AZ1.Drive not ready
        [11].rgxStoppingFaults[0].4   // A69AZ1.Drive not ready
        [12].rgxStoppingFaults[0].4   // A70AZ1.Drive not ready
        [13].rgxStoppingFaults[0].4   // A71AZ1.Drive not ready
        [14].rgxStoppingFaults[0].4   // A72AZ1.Drive not ready
        [15].rgxStoppingFaults[0].4   // A73AZ1.Drive not ready
        [16].rgxStoppingFaults[0].4   // A74AZ1.Drive not ready
        [17].rgxStoppingFaults[0].4   // A77AZ1.Drive not ready
        [18].rgxStoppingFaults[0].4   // A75AZ1.Drive not ready
        [19].rgxStoppingFaults[0].4   // A76AZ1.Drive not ready
   M2xx_CONVEYOR_HMR : MAC_CONVEYOR_HMR[20] := ([0].dStatus := 1, [1].dStatus := 1, [2].dStatus := 1, [3].dStatus := 1, [4].dStatus := 1, [5].dStatus := 7, [6].dStatus := 7, [7].dStatus := 7, [8].dStatus := 7, [9].dStatus := 7, [10].dStatus := 7, [11].dStatus := 1, [12].dStatus := 1, [13].dStatus := 1, [14].dStatus := 1, [15].dStatus := 1, [16].dStatus := 1, [17].dStatus := 1, [18].dStatus := 1, [19].dStatus := 1); {access Read Only}
        [0]   // M202
        [10]   // M213
        [11]   // M214
        [1]   // M203
        [2]   // M204
        [3]   // M206
        [4]   // M207
        [5]   // M208
        [6]   // M209
        [7]   // M210
        [8]   // M211
        [9]   // M212
        [17]   // M220
        [16]   // M219
        [15]   // M218
        [18]   // M301M1
        [14]   // M217
        [13]   // M216
        [12]   // M215
        [19]   // M301M2
   M2xx_CONVEYOR_HMW : MAC_CONVEYOR_HMW[20];
        [0]   // M202
        [10]   // M213
        [11]   // M214
        [1]   // M203
        [2]   // M204
        [3]   // M206
        [4]   // M207
        [5]   // M208
        [6]   // M209
        [7]   // M210
        [8]   // M211
        [9]   // M212
        [18]   // M301M1
        [17]   // M220
        [16]   // M219
        [15]   // M218
        [14]   // M217
        [13]   // M216
        [12]   // M215
        [19]   // M301M2
   M2xx_CONVEYOR_IN_MOTION : MAC_CONVEYOR_IN_MOTION[20]; {access None}
   M2xx_CONVEYOR_OUT_MOTION : MAC_CONVEYOR_OUT_MOTION[20] := ([0].DR_MSO_M.FLAGS := 33554432, [0].DR_MSF_M.FLAGS := -1577058304, [0].DR_MSF_M.EN := 1, [0].DR_MSF_M.DN := 1, [0].DR_MSF_M.STATUS := 2, [0].DR_MSF_M.STATE := 1, [0].DR_MASR_M.FLAGS := 33554432, [0].DR_MAJ_M.FLAGS := 33554432, [0].DR_MCD_M.FLAGS := 33554432, [0].DR_MAS_M.FLAGS := -1442840576, [0].DR_MAS_M.EN := 1, [0].DR_MAS_M.DN := 1, [0].DR_MAS_M.PC := 1, [1].DR_MSO_M.FLAGS := 33554432, [1].DR_MSF_M.FLAGS := -1577058304, [1].DR_MSF_M.EN := 1, [1].DR_MSF_M.DN := 1, [1].DR_MSF_M.STATUS := 2, [1].DR_MSF_M.STATE := 1, [1].DR_MASR_M.FLAGS := 33554432, [1].DR_MAJ_M.FLAGS := 33554432, [1].DR_MCD_M.FLAGS := 33554432, [1].DR_MAS_M.FLAGS := -1442840576, [1].DR_MAS_M.EN := 1, [1].DR_MAS_M.DN := 1, [1].DR_MAS_M.PC := 1, [2].DR_MSO_M.FLAGS := 33554432, [2].DR_MSF_M.FLAGS := -1577058304, [2].DR_MSF_M.EN := 1, [2].DR_MSF_M.DN := 1, [2].DR_MSF_M.STATUS := 2, [2].DR_MSF_M.STATE := 1, [2].DR_MASR_M.FLAGS := 33554432, [2].DR_MAJ_M.FLAGS := 33554432, [2].DR_MCD_M.FLAGS := 33554432, [2].DR_MAS_M.FLAGS := -1442840576, [2].DR_MAS_M.EN := 1, [2].DR_MAS_M.DN := 1, [2].DR_MAS_M.PC := 1, [3].DR_MSO_M.FLAGS := 33554432, [3].DR_MSF_M.FLAGS := -1577058304, [3].DR_MSF_M.EN := 1, [3].DR_MSF_M.DN := 1, [3].DR_MSF_M.STATUS := 2, [3].DR_MSF_M.STATE := 1, [3].DR_MASR_M.FLAGS := 33554432, [3].DR_MAJ_M.FLAGS := 33554432, [3].DR_MCD_M.FLAGS := 33554432, [3].DR_MAS_M.FLAGS := -1442840576, [3].DR_MAS_M.EN := 1, [3].DR_MAS_M.DN := 1, [3].DR_MAS_M.PC := 1, [4].DR_MSO_M.FLAGS := 33554432, [4].DR_MSF_M.FLAGS := -1577058304, [4].DR_MSF_M.EN := 1, [4].DR_MSF_M.DN := 1, [4].DR_MSF_M.STATUS := 2, [4].DR_MSF_M.STATE := 1, [4].DR_MASR_M.FLAGS := 33554432, [4].DR_MAJ_M.FLAGS := 33554432,
        [4].DR_MCD_M.FLAGS := 33554432, [4].DR_MAS_M.FLAGS := -1442840576, [4].DR_MAS_M.EN := 1, [4].DR_MAS_M.DN := 1, [4].DR_MAS_M.PC := 1, [5].DR_MSO_M.FLAGS := 33554432, [5].DR_MSF_M.FLAGS := -1577058304, [5].DR_MSF_M.EN := 1, [5].DR_MSF_M.DN := 1, [5].DR_MSF_M.STATUS := 2, [5].DR_MSF_M.STATE := 1, [5].DR_MASR_M.FLAGS := 33554432, [5].DR_MAJ_M.FLAGS := 33554432, [5].DR_MCD_M.FLAGS := 33554432, [5].DR_MAS_M.FLAGS := -1442840576, [5].DR_MAS_M.EN := 1, [5].DR_MAS_M.DN := 1, [5].DR_MAS_M.PC := 1, [6].DR_MSO_M.FLAGS := 33554432, [6].DR_MSF_M.FLAGS := -1577058304, [6].DR_MSF_M.EN := 1, [6].DR_MSF_M.DN := 1, [6].DR_MSF_M.STATUS := 2, [6].DR_MSF_M.STATE := 1, [6].DR_MASR_M.FLAGS := 33554432, [6].DR_MAJ_M.FLAGS := 33554432, [6].DR_MCD_M.FLAGS := 33554432, [6].DR_MAS_M.FLAGS := -1442840576, [6].DR_MAS_M.EN := 1, [6].DR_MAS_M.DN := 1, [6].DR_MAS_M.PC := 1, [7].DR_MSO_M.FLAGS := 33554432, [7].DR_MSF_M.FLAGS := -1577058304, [7].DR_MSF_M.EN := 1, [7].DR_MSF_M.DN := 1, [7].DR_MSF_M.STATUS := 2, [7].DR_MSF_M.STATE := 1, [7].DR_MASR_M.FLAGS := 33554432, [7].DR_MAJ_M.FLAGS := 33554432, [7].DR_MCD_M.FLAGS := 33554432, [7].DR_MAS_M.FLAGS := -1442840576, [7].DR_MAS_M.EN := 1, [7].DR_MAS_M.DN := 1, [7].DR_MAS_M.PC := 1, [8].DR_MSO_M.FLAGS := 33554432, [8].DR_MSF_M.FLAGS := -1577058304, [8].DR_MSF_M.EN := 1, [8].DR_MSF_M.DN := 1, [8].DR_MSF_M.STATUS := 2, [8].DR_MSF_M.STATE := 1, [8].DR_MASR_M.FLAGS := 33554432, [8].DR_MAJ_M.FLAGS := 33554432, [8].DR_MCD_M.FLAGS := 33554432, [8].DR_MAS_M.FLAGS := -1442840576, [8].DR_MAS_M.EN := 1, [8].DR_MAS_M.DN := 1, [8].DR_MAS_M.PC := 1, [9].DR_MSO_M.FLAGS := 33554432, [9].DR_MSF_M.FLAGS := -1577058304, [9].DR_MSF_M.EN := 1,
        [9].DR_MSF_M.DN := 1, [9].DR_MSF_M.STATUS := 2, [9].DR_MSF_M.STATE := 1, [9].DR_MASR_M.FLAGS := 33554432, [9].DR_MAJ_M.FLAGS := 33554432, [9].DR_MCD_M.FLAGS := 33554432, [9].DR_MAS_M.FLAGS := -1442840576, [9].DR_MAS_M.EN := 1, [9].DR_MAS_M.DN := 1, [9].DR_MAS_M.PC := 1, [10].DR_MSO_M.FLAGS := 33554432, [10].DR_MSF_M.FLAGS := -1577058304, [10].DR_MSF_M.EN := 1, [10].DR_MSF_M.DN := 1, [10].DR_MSF_M.STATUS := 2, [10].DR_MSF_M.STATE := 1, [10].DR_MASR_M.FLAGS := 33554432, [10].DR_MAJ_M.FLAGS := 33554432, [10].DR_MCD_M.FLAGS := 33554432, [10].DR_MAS_M.FLAGS := -1442840576, [10].DR_MAS_M.EN := 1, [10].DR_MAS_M.DN := 1, [10].DR_MAS_M.PC := 1, [11].DR_MSO_M.FLAGS := 33554432, [11].DR_MSF_M.FLAGS := -1577058304, [11].DR_MSF_M.EN := 1, [11].DR_MSF_M.DN := 1, [11].DR_MSF_M.STATUS := 2, [11].DR_MSF_M.STATE := 1, [11].DR_MASR_M.FLAGS := 33554432, [11].DR_MAJ_M.FLAGS := 33554432, [11].DR_MCD_M.FLAGS := 33554432, [11].DR_MAS_M.FLAGS := -1442840576, [11].DR_MAS_M.EN := 1, [11].DR_MAS_M.DN := 1, [11].DR_MAS_M.PC := 1, [12].DR_MSO_M.FLAGS := 33554432, [12].DR_MSF_M.FLAGS := -1577058304, [12].DR_MSF_M.EN := 1, [12].DR_MSF_M.DN := 1, [12].DR_MSF_M.STATUS := 2, [12].DR_MSF_M.STATE := 1, [12].DR_MASR_M.FLAGS := 33554432, [12].DR_MAJ_M.FLAGS := 33554432, [12].DR_MCD_M.FLAGS := 33554432, [12].DR_MAS_M.FLAGS := -1845493760, [12].DR_MAS_M.EN := 1, [12].DR_MAS_M.ER := 1, [12].DR_MAS_M.ERR := 13, [12].DR_MAS_M.EXERR := 4, [13].DR_MSO_M.FLAGS := 33554432, [13].DR_MSF_M.FLAGS := -1577058304, [13].DR_MSF_M.EN := 1, [13].DR_MSF_M.DN := 1, [13].DR_MSF_M.STATUS := 2, [13].DR_MSF_M.STATE := 1, [13].DR_MASR_M.FLAGS := 33554432, [13].DR_MAJ_M.FLAGS := 33554432, [13].DR_MCD_M.FLAGS := 33554432, [13].DR_MAS_M.FLAGS := -1845493760,
        [13].DR_MAS_M.EN := 1, [13].DR_MAS_M.ER := 1, [13].DR_MAS_M.ERR := 13, [13].DR_MAS_M.EXERR := 4, [14].DR_MSO_M.FLAGS := 33554432, [14].DR_MSF_M.FLAGS := -1577058304, [14].DR_MSF_M.EN := 1, [14].DR_MSF_M.DN := 1, [14].DR_MSF_M.STATUS := 2, [14].DR_MSF_M.STATE := 1, [14].DR_MASR_M.FLAGS := 33554432, [14].DR_MAJ_M.FLAGS := 33554432, [14].DR_MCD_M.FLAGS := 33554432, [14].DR_MAS_M.FLAGS := -1845493760, [14].DR_MAS_M.EN := 1, [14].DR_MAS_M.ER := 1, [14].DR_MAS_M.ERR := 13, [14].DR_MAS_M.EXERR := 4, [15].DR_MSO_M.FLAGS := 33554432, [15].DR_MSF_M.FLAGS := -1577058304, [15].DR_MSF_M.EN := 1, [15].DR_MSF_M.DN := 1, [15].DR_MSF_M.STATUS := 2, [15].DR_MSF_M.STATE := 1, [15].DR_MASR_M.FLAGS := 33554432, [15].DR_MAJ_M.FLAGS := 33554432, [15].DR_MCD_M.FLAGS := 33554432, [15].DR_MAS_M.FLAGS := -1845493760, [15].DR_MAS_M.EN := 1, [15].DR_MAS_M.ER := 1, [15].DR_MAS_M.ERR := 13, [15].DR_MAS_M.EXERR := 4, [16].DR_MSO_M.FLAGS := 33554432, [16].DR_MSF_M.FLAGS := -1577058304, [16].DR_MSF_M.EN := 1, [16].DR_MSF_M.DN := 1, [16].DR_MSF_M.STATUS := 2, [16].DR_MSF_M.STATE := 1, [16].DR_MASR_M.FLAGS := 33554432, [16].DR_MAJ_M.FLAGS := 33554432, [16].DR_MCD_M.FLAGS := 33554432, [16].DR_MAS_M.FLAGS := -1845493760, [16].DR_MAS_M.EN := 1, [16].DR_MAS_M.ER := 1, [16].DR_MAS_M.ERR := 13, [16].DR_MAS_M.EXERR := 4, [17].DR_MSO_M.FLAGS := 33554432, [17].DR_MSF_M.FLAGS := -1577058304, [17].DR_MSF_M.EN := 1, [17].DR_MSF_M.DN := 1, [17].DR_MSF_M.STATUS := 2, [17].DR_MSF_M.STATE := 1, [17].DR_MASR_M.FLAGS := 33554432, [17].DR_MAJ_M.FLAGS := 33554432, [17].DR_MCD_M.FLAGS := 33554432, [17].DR_MAS_M.FLAGS := -1845493760, [17].DR_MAS_M.EN := 1, [17].DR_MAS_M.ER := 1, [17].DR_MAS_M.ERR := 13, [17].DR_MAS_M.EXERR := 4,
        [18].DR_MSO_M.FLAGS := 33554432, [18].DR_MSF_M.FLAGS := -1577058304, [18].DR_MSF_M.EN := 1, [18].DR_MSF_M.DN := 1, [18].DR_MSF_M.STATUS := 2, [18].DR_MSF_M.STATE := 1, [18].DR_MASR_M.FLAGS := 33554432, [18].DR_MAJ_M.FLAGS := 33554432, [18].DR_MCD_M.FLAGS := 33554432, [18].DR_MAS_M.FLAGS := -1845493760, [18].DR_MAS_M.EN := 1, [18].DR_MAS_M.ER := 1, [18].DR_MAS_M.ERR := 13, [18].DR_MAS_M.EXERR := 4, [19].DR_MSO_M.FLAGS := 33554432, [19].DR_MSF_M.FLAGS := -1577058304, [19].DR_MSF_M.EN := 1, [19].DR_MSF_M.DN := 1, [19].DR_MSF_M.STATUS := 2, [19].DR_MSF_M.STATE := 1, [19].DR_MASR_M.FLAGS := 33554432, [19].DR_MAJ_M.FLAGS := 33554432, [19].DR_MCD_M.FLAGS := 33554432, [19].DR_MAS_M.FLAGS := -1845493760, [19].DR_MAS_M.EN := 1, [19].DR_MAS_M.ER := 1, [19].DR_MAS_M.ERR := 13, [19].DR_MAS_M.EXERR := 4); {access None}
   M301_M1_DR : AXIS_CIP_DRIVE; {access Read Only}
   M301_M1_DR_IN_MAJ : MOTION_INSTRUCTION := (FLAGS := 570425344, DN := 1); {access None}
   M301_M1_DR_IN_MAM : MOTION_INSTRUCTION := (FLAGS := 33554432); {access None}
   M301_M1_DR_IN_MAR : MOTION_INSTRUCTION := (FLAGS := 33554432); {access None}
   M301_M1_DR_IN_MAS : MOTION_INSTRUCTION := (FLAGS := -1442840576, EN := 1, DN := 1, PC := 1); {access None}
   M301_M1_DR_IN_MCD : MOTION_INSTRUCTION := (FLAGS := 570425344, DN := 1); {access None}
   M301_M1_DR_IN_MRP : MOTION_INSTRUCTION := (FLAGS := 33554432); {access None}
   M301_M1_DR_MAFR : MOTION_INSTRUCTION := (FLAGS := 301989888, ER := 1, ERR := 11); {access None}
   M301_M1_DR_MDR : MOTION_INSTRUCTION := (FLAGS := -1845493760, EN := 1, ER := 1, ERR := 11); {access None}
   M301_M1_DR_MSF : MOTION_INSTRUCTION := (FLAGS := 570425344, DN := 1, STATUS := 2, STATE := 1); {access None}
   M301_M1_DR_MSO : MOTION_INSTRUCTION := (FLAGS := -1610612736, EN := 1, DN := 1, STATE := 1); {access None}
   M301_M1_DR_OUT_MAJ : MOTION_INSTRUCTION := (FLAGS := 570425344, DN := 1); {access None}
   M301_M1_DR_OUT_MAM : MOTION_INSTRUCTION := (FLAGS := 33554432); {access None}
   M301_M1_DR_OUT_MAR : MOTION_INSTRUCTION := (FLAGS := 33554432); {access None}
   M301_M1_DR_OUT_MAS : MOTION_INSTRUCTION := (FLAGS := -1442840576, EN := 1, DN := 1, PC := 1); {access None}
   M301_M1_DR_OUT_MCD : MOTION_INSTRUCTION := (FLAGS := 570425344, DN := 1); {access None}
   M301_M1_DR_OUT_MRP : MOTION_INSTRUCTION := (FLAGS := 33554432); {access None}
   M301_M2_DR : AXIS_CIP_DRIVE; {access Read Only}
   M301_M2_DR_IN_MAJ : MOTION_INSTRUCTION := (FLAGS := 570425344, DN := 1); {access None}
   M301_M2_DR_IN_MAM : MOTION_INSTRUCTION := (FLAGS := 33554432); {access None}
   M301_M2_DR_IN_MAR : MOTION_INSTRUCTION := (FLAGS := 33554432); {access None}
   M301_M2_DR_IN_MAS : MOTION_INSTRUCTION := (FLAGS := -1442840576, EN := 1, DN := 1, PC := 1); {access None}
   M301_M2_DR_IN_MCD : MOTION_INSTRUCTION := (FLAGS := 570425344, DN := 1); {access None}
   M301_M2_DR_IN_MRP : MOTION_INSTRUCTION := (FLAGS := 33554432); {access None}
   M301_M2_DR_MAFR : MOTION_INSTRUCTION := (FLAGS := 301989888, ER := 1, ERR := 11); {access None}
   M301_M2_DR_MDR : MOTION_INSTRUCTION := (FLAGS := -1845493760, EN := 1, ER := 1, ERR := 11); {access None}
   M301_M2_DR_MSF : MOTION_INSTRUCTION := (FLAGS := 570425344, DN := 1, STATUS := 2, STATE := 1); {access None}
   M301_M2_DR_MSO : MOTION_INSTRUCTION := (FLAGS := -1610612736, EN := 1, DN := 1, STATE := 1); {access None}
   M301_M2_DR_OUT_MAJ : MOTION_INSTRUCTION := (FLAGS := 570425344, DN := 1); {access None}
   M301_M2_DR_OUT_MAM : MOTION_INSTRUCTION := (FLAGS := 33554432); {access None}
   M301_M2_DR_OUT_MAR : MOTION_INSTRUCTION := (FLAGS := 33554432); {access None}
   M301_M2_DR_OUT_MAS : MOTION_INSTRUCTION := (FLAGS := -1442840576, EN := 1, DN := 1, PC := 1); {access None}
   M301_M2_DR_OUT_MCD : MOTION_INSTRUCTION := (FLAGS := 570425344, DN := 1); {access None}
   M301_M2_DR_OUT_MRP : MOTION_INSTRUCTION := (FLAGS := 33554432); {access None}
   M32_MMI : ALIAS FOR N54[376].3;
   M37B_FWD_DIR : ALIAS FOR B3[1].14;
   M37B_FWD_PL : ALIAS FOR O[25].5;
   M37B_FWD_SIG : ALIAS FOR I[112].3;
   M37B_FWD_SS : ALIAS FOR I[24].8;
   M37B_REV_DIR : ALIAS FOR B3[1].15;
   M37B_REV_PL : ALIAS FOR O[25].6;
   M37B_REV_SIG : ALIAS FOR I[112].4;
   M37B_REV_SS : ALIAS FOR I[24].9;
   M37B_RUN_FWD : ALIAS FOR O[119].0;
   M37B_RUN_REV : ALIAS FOR O[119].1;
   M40_MMI : ALIAS FOR N54[376].1;
   M41_MMI : ALIAS FOR N54[375].15;
   M42_MMI : ALIAS FOR N54[376].0;
   M43_MMI : ALIAS FOR N54[375].14;
   M47_REV_SS : ALIAS FOR I[24].11;
   M47B_FWD_DIR : ALIAS FOR B3[1].12;
   M47B_FWD_PL : ALIAS FOR O[25].7;
   M47B_FWD_SIG : ALIAS FOR I[112].1;
   M47B_FWD_SS : ALIAS FOR I[24].10;
   M47B_REV_DIR : ALIAS FOR B3[1].13;
   M47B_REV_PL : ALIAS FOR O[25].8;
   M47B_REV_SIG : ALIAS FOR I[112].2;
   M47B_REV_SS : ALIAS FOR I[1].8;
   M47B_RUN_FWD : ALIAS FOR O[119].2;
   M47B_RUN_REV : ALIAS FOR O[119].3;
   MADSEN_2IN_PULS : ALIAS FOR I[12].15;
   MB_ALM_RESET : ALIAS FOR I[16].10;